REGION Network 10: Bit 9
   RUNG wire#powerrail
      Contact( #wInWord.%X9 )
      Coil( #bOutBit09 )
   END_RUNG
   // the same network as SCL:
   #bOutBit09 := #wInWord.%X9;
END_REGION

REGION Network 11: Bit 10
   RUNG wire#powerrail
      Contact( #wInWord.%X10 )
      Coil( #bOutBit10 )
   END_RUNG
   // the same network as SCL:
   #bOutBit10 := #wInWord.%X10;
END_REGION

REGION Network 12: Bit 11
   RUNG wire#powerrail
      Contact( #wInWord.%X11 )
      Coil( #bOutBit11 )
   END_RUNG
   // the same network as SCL:
   #bOutBit11 := #wInWord.%X11;
END_REGION

REGION Network 13: Bit 12
   RUNG wire#powerrail
      Contact( #wInWord.%X12 )
      Coil( #bOutBit12 )
   END_RUNG
   // the same network as SCL:
   #bOutBit12 := #wInWord.%X12;
END_REGION

REGION Network 14: Bit 13
   RUNG wire#powerrail
      Contact( #wInWord.%X13 )
      Coil( #bOutBit13 )
   END_RUNG
   // the same network as SCL:
   #bOutBit13 := #wInWord.%X13;
END_REGION

REGION Network 15: Bit 14
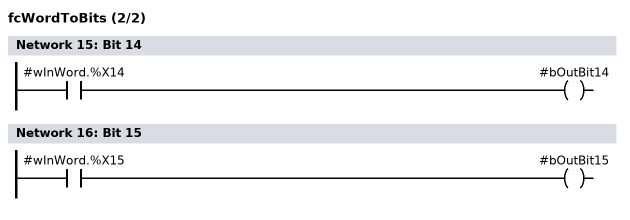
   RUNG wire#powerrail
      Contact( #wInWord.%X14 )
      Coil( #bOutBit14 )
   END_RUNG
   // the same network as SCL:
   #bOutBit14 := #wInWord.%X14;
END_REGION

REGION Network 16: Bit 15
   RUNG wire#powerrail
      Contact( #wInWord.%X15 )
      Coil( #bOutBit15 )
   END_RUNG
   // the same network as SCL:
   #bOutBit15 := #wInWord.%X15;
END_REGION
END_FUNCTION

FUNCTION "fcBitsToWord" : Void   // FC1001, LAD
TITLE = Pack Bits into word
{ S7_Optimized_Access := 'FALSE' }
AUTHOR : DMC
FAMILY : LowLevel
VERSION : 0.1
BEGIN

REGION Network 1: Bit0
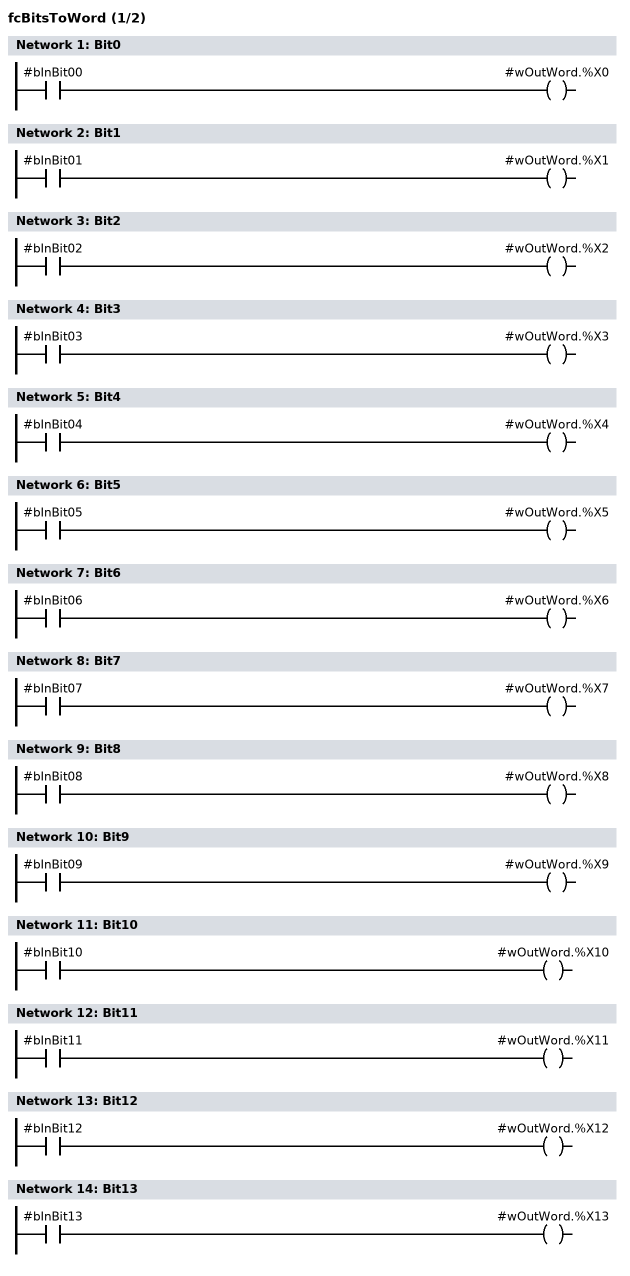
   RUNG wire#powerrail
      Contact( #bInBit00 )
      Coil( #wOutWord.%X0 )
   END_RUNG
   // the same network as SCL:
   #wOutWord.%X0 := #bInBit00;
END_REGION

REGION Network 2: Bit1
   RUNG wire#powerrail
      Contact( #bInBit01 )
      Coil( #wOutWord.%X1 )
   END_RUNG
   // the same network as SCL:
   #wOutWord.%X1 := #bInBit01;
END_REGION

REGION Network 3: Bit2
   RUNG wire#powerrail
      Contact( #bInBit02 )
      Coil( #wOutWord.%X2 )
   END_RUNG
   // the same network as SCL:
   #wOutWord.%X2 := #bInBit02;
END_REGION

REGION Network 4: Bit3
   RUNG wire#powerrail
      Contact( #bInBit03 )
      Coil( #wOutWord.%X3 )
   END_RUNG
   // the same network as SCL:
   #wOutWord.%X3 := #bInBit03;
END_REGION

REGION Network 5: Bit4
   RUNG wire#powerrail
      Contact( #bInBit04 )
      Coil( #wOutWord.%X4 )
   END_RUNG
   // the same network as SCL:
   #wOutWord.%X4 := #bInBit04;
END_REGION

REGION Network 6: Bit5
   RUNG wire#powerrail
      Contact( #bInBit05 )
      Coil( #wOutWord.%X5 )
   END_RUNG
   // the same network as SCL:
   #wOutWord.%X5 := #bInBit05;
END_REGION

REGION Network 7: Bit6
   RUNG wire#powerrail
      Contact( #bInBit06 )
      Coil( #wOutWord.%X6 )
   END_RUNG
   // the same network as SCL:
   #wOutWord.%X6 := #bInBit06;
END_REGION

REGION Network 8: Bit7
   RUNG wire#powerrail
      Contact( #bInBit07 )
      Coil( #wOutWord.%X7 )
   END_RUNG
   // the same network as SCL:
   #wOutWord.%X7 := #bInBit07;
END_REGION

REGION Network 9: Bit8
   RUNG wire#powerrail
      Contact( #bInBit08 )
      Coil( #wOutWord.%X8 )
   END_RUNG
   // the same network as SCL:
   #wOutWord.%X8 := #bInBit08;
END_REGION

REGION Network 10: Bit9
   RUNG wire#powerrail
      Contact( #bInBit09 )
      Coil( #wOutWord.%X9 )
   END_RUNG
   // the same network as SCL:
   #wOutWord.%X9 := #bInBit09;
END_REGION

REGION Network 11: Bit10
   RUNG wire#powerrail
      Contact( #bInBit10 )
      Coil( #wOutWord.%X10 )
   END_RUNG
   // the same network as SCL:
   #wOutWord.%X10 := #bInBit10;
END_REGION

REGION Network 12: Bit11
   RUNG wire#powerrail
      Contact( #bInBit11 )
      Coil( #wOutWord.%X11 )
   END_RUNG
   // the same network as SCL:
   #wOutWord.%X11 := #bInBit11;
END_REGION

REGION Network 13: Bit12
   RUNG wire#powerrail
      Contact( #bInBit12 )
      Coil( #wOutWord.%X12 )
   END_RUNG
   // the same network as SCL:
   #wOutWord.%X12 := #bInBit12;
END_REGION

REGION Network 14: Bit13
   RUNG wire#powerrail
      Contact( #bInBit13 )
      Coil( #wOutWord.%X13 )
   END_RUNG
   // the same network as SCL:
   #wOutWord.%X13 := #bInBit13;
END_REGION

REGION Network 15: Bit14
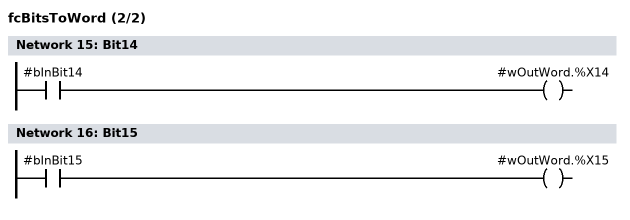
   RUNG wire#powerrail
      Contact( #bInBit14 )
      Coil( #wOutWord.%X14 )
   END_RUNG
   // the same network as SCL:
   #wOutWord.%X14 := #bInBit14;
END_REGION

REGION Network 16: Bit15
   RUNG wire#powerrail
      Contact( #bInBit15 )
      Coil( #wOutWord.%X15 )
   END_RUNG
   // the same network as SCL:
   #wOutWord.%X15 := #bInBit15;
END_REGION
END_FUNCTION

// folder: Library Blocks/Resources/HMI

FUNCTION_BLOCK "fbErrorScroller"   // FB1007, LAD
TITLE = Scrolls through the error codes for display on the HMI
{ S7_Optimized_Access := 'FALSE' }
AUTHOR : DMC
FAMILY : Error
VERSION : 0.1
   VAR_TEMP   // added for the SCL form of the ladder/FBD networks
      _w1 : Bool;
   END_VAR
BEGIN

REGION Network 1: Error Exists
   // OR all of the possible errors. If any error Exists, SET bErrorExists
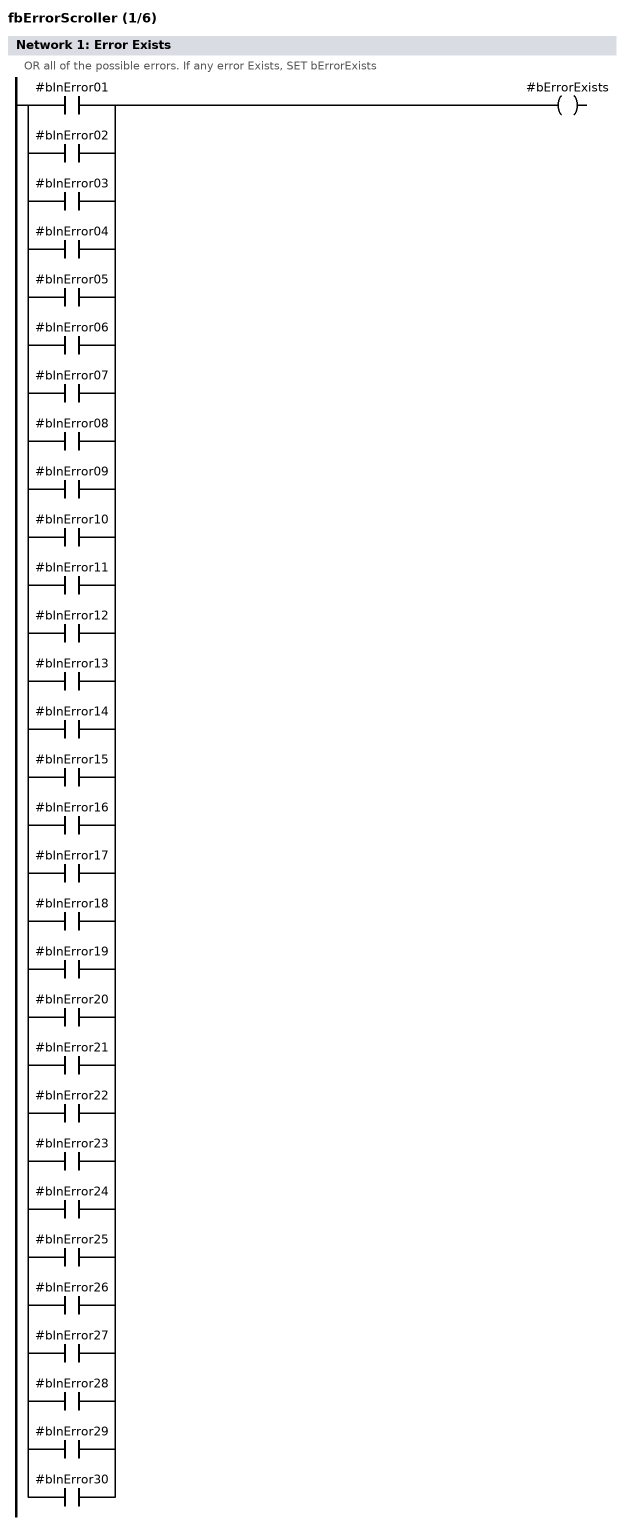
   RUNG wire#powerrail
      Contact( #bInError01 )
      wire#w1
      Coil( #bErrorExists )
   END_RUNG
   RUNG wire#powerrail
      Contact( #bInError02 )
   END_RUNG wire#w1
   RUNG wire#powerrail
      Contact( #bInError03 )
   END_RUNG wire#w1
   RUNG wire#powerrail
      Contact( #bInError04 )
   END_RUNG wire#w1
   RUNG wire#powerrail
      Contact( #bInError05 )
   END_RUNG wire#w1
   RUNG wire#powerrail
      Contact( #bInError06 )
   END_RUNG wire#w1
   RUNG wire#powerrail
      Contact( #bInError07 )
   END_RUNG wire#w1
   RUNG wire#powerrail
      Contact( #bInError08 )
   END_RUNG wire#w1
   RUNG wire#powerrail
      Contact( #bInError09 )
   END_RUNG wire#w1
   RUNG wire#powerrail
      Contact( #bInError10 )
   END_RUNG wire#w1
   RUNG wire#powerrail
      Contact( #bInError11 )
   END_RUNG wire#w1
   RUNG wire#powerrail
      Contact( #bInError12 )
   END_RUNG wire#w1
   RUNG wire#powerrail
      Contact( #bInError13 )
   END_RUNG wire#w1
   RUNG wire#powerrail
      Contact( #bInError14 )
   END_RUNG wire#w1
   RUNG wire#powerrail
      Contact( #bInError15 )
   END_RUNG wire#w1
   RUNG wire#powerrail
      Contact( #bInError16 )
   END_RUNG wire#w1
   RUNG wire#powerrail
      Contact( #bInError17 )
   END_RUNG wire#w1
   RUNG wire#powerrail
      Contact( #bInError18 )
   END_RUNG wire#w1
   RUNG wire#powerrail
      Contact( #bInError19 )
   END_RUNG wire#w1
   RUNG wire#powerrail
      Contact( #bInError20 )
   END_RUNG wire#w1
   RUNG wire#powerrail
      Contact( #bInError21 )
   END_RUNG wire#w1
   RUNG wire#powerrail
      Contact( #bInError22 )
   END_RUNG wire#w1
   RUNG wire#powerrail
      Contact( #bInError23 )
   END_RUNG wire#w1
   RUNG wire#powerrail
      Contact( #bInError24 )
   END_RUNG wire#w1
   RUNG wire#powerrail
      Contact( #bInError25 )
   END_RUNG wire#w1
   RUNG wire#powerrail
      Contact( #bInError26 )
   END_RUNG wire#w1
   RUNG wire#powerrail
      Contact( #bInError27 )
   END_RUNG wire#w1
   RUNG wire#powerrail
      Contact( #bInError28 )
   END_RUNG wire#w1
   RUNG wire#powerrail
      Contact( #bInError29 )
   END_RUNG wire#w1
   RUNG wire#powerrail
      Contact( #bInError30 )
   END_RUNG wire#w1
   // the same network as SCL:
   #bErrorExists := #bInError01 OR #bInError02 OR #bInError03 OR #bInError04 OR #bInError05 OR #bInError06 OR #bInError07 OR #bInError08 OR #bInError09 OR #bInError10 OR #bInError11 OR #bInError12 OR #bInError13 OR #bInError14 OR #bInError15 OR #bInError16 OR #bInError17 OR #bInError18 OR #bInError19 OR #bInError20 OR #bInError21 OR #bInError22 OR #bInError23 OR #bInError24 OR #bInError25 OR #bInError26 OR #bInError27 OR #bInError28 OR #bInError29 OR #bInError30;
END_REGION

REGION Network 2
   // ============================ Scroll errors on HMI ========================
   // Timed delay
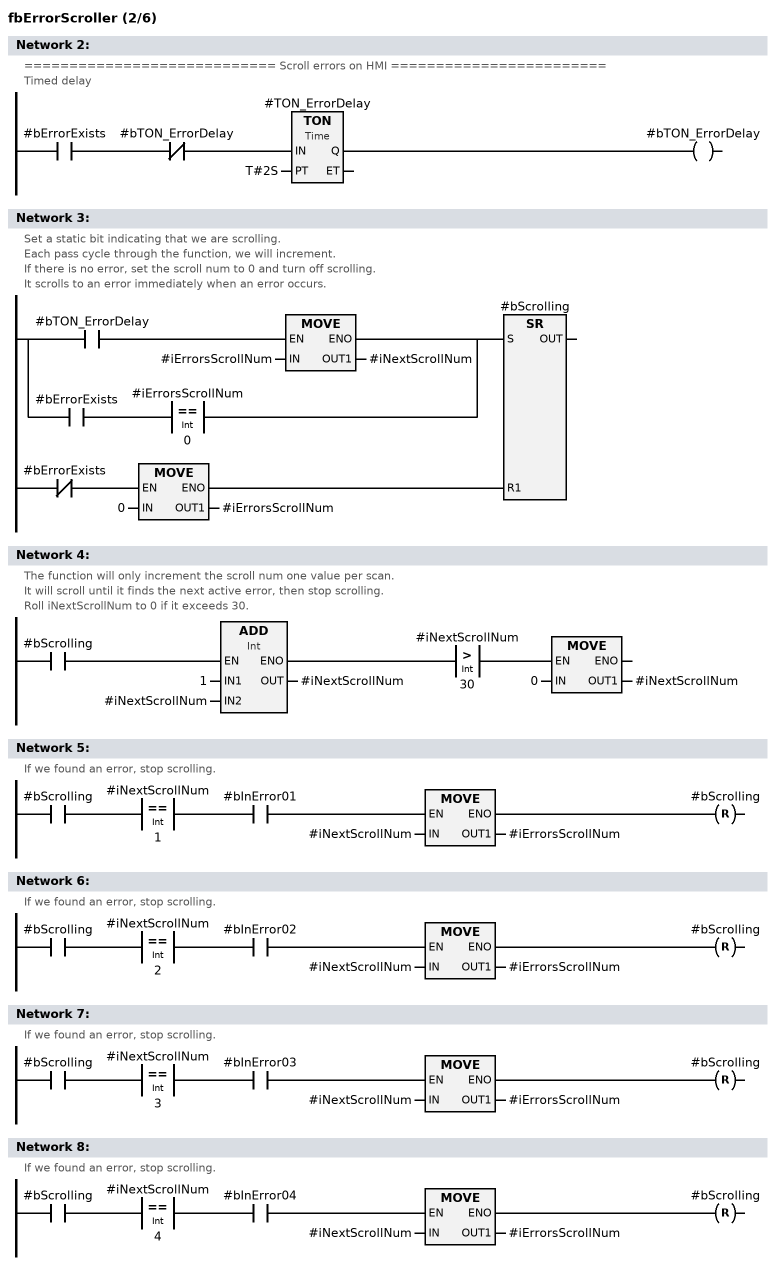
   #TON_ErrorDelay.TON(IN := #bErrorExists AND NOT #bTON_ErrorDelay, PT := T#2S);
   #bTON_ErrorDelay := #TON_ErrorDelay.Q;
END_REGION

REGION Network 3
   // Set a static bit indicating that we are scrolling.  
   // Each pass cycle through the function, we will increment.  
   // If there is no error, set the scroll num to 0 and turn off scrolling.  
   // It scrolls to an error immediately when an error occurs.
   RUNG wire#powerrail
      Contact( #bTON_ErrorDelay )
      { S7_GenerateENO := "TRUE" } Move(in := #iErrorsScrollNum, out1 => #iNextScrollNum)
      wire#w1
      S_SR(operand := #bScrolling, r1 := wire#w2)
   END_RUNG
   RUNG wire#powerrail
      Contact( #bErrorExists )
      { S7_Templates := "SrcType := Int" } EQ_Contact(in1 := #iErrorsScrollNum, in2 := 0)
   END_RUNG wire#w1
   RUNG wire#powerrail
      I_Contact( #bErrorExists )
      { S7_GenerateENO := "TRUE" } Move(in := 0, out1 => #iErrorsScrollNum)
   END_RUNG wire#w2
   // the same network as SCL:
   // ENO of a box is taken as its EN; it also drops when the box reports an error
   IF #bTON_ErrorDelay THEN #iNextScrollNum := #iErrorsScrollNum; END_IF;
   #_w1 := #bTON_ErrorDelay OR (#bErrorExists AND (#iErrorsScrollNum = 0));
   IF NOT #bErrorExists THEN #iErrorsScrollNum := 0; END_IF;
   IF #_w1 THEN
       #bScrolling := TRUE;   // SR flip-flop
   END_IF;
   IF NOT #bErrorExists THEN #bScrolling := FALSE; END_IF;
END_REGION

REGION Network 4
   // The function will only increment the scroll num one value per scan.  
   // It will scroll until it finds the next active error, then stop scrolling.  
   // Roll iNextScrollNum to 0 if it exceeds 30.
   RUNG wire#powerrail
      Contact( #bScrolling )
      { S7_Templates := "SrcType := Int"; S7_GenerateENO := "TRUE" } Add(in1 := 1, in2 := #iNextScrollNum, out => #iNextScrollNum)
      { S7_Templates := "SrcType := Int" } GT_Contact(in1 := #iNextScrollNum, in2 := 30)
      { S7_GenerateENO := "TRUE" } Move(in := 0, out1 => #iNextScrollNum)
   END_RUNG
   // the same network as SCL:
   // ENO of a box is taken as its EN; it also drops when the box reports an error
   IF #bScrolling THEN #iNextScrollNum := 1 + #iNextScrollNum; END_IF;
   IF #bScrolling AND (#iNextScrollNum > 30) THEN #iNextScrollNum := 0; END_IF;
END_REGION

REGION Network 5
   // If we found an error, stop scrolling.
   RUNG wire#powerrail
      Contact( #bScrolling )
      { S7_Templates := "SrcType := Int" } EQ_Contact(in1 := #iNextScrollNum, in2 := 1)
      Contact( #bInError01 )
      { S7_GenerateENO := "TRUE" } Move(in := #iNextScrollNum, out1 => #iErrorsScrollNum)
      R_Coil( #bScrolling )
   END_RUNG
   // the same network as SCL:
   // ENO of a box is taken as its EN; it also drops when the box reports an error
   IF #bScrolling AND (#iNextScrollNum = 1) AND #bInError01 THEN
       #iErrorsScrollNum := #iNextScrollNum;
       #bScrolling := FALSE;
   END_IF;
END_REGION

REGION Network 6
   // If we found an error, stop scrolling.
   RUNG wire#powerrail
      Contact( #bScrolling )
      { S7_Templates := "SrcType := Int" } EQ_Contact(in1 := #iNextScrollNum, in2 := 2)
      Contact( #bInError02 )
      { S7_GenerateENO := "TRUE" } Move(in := #iNextScrollNum, out1 => #iErrorsScrollNum)
      R_Coil( #bScrolling )
   END_RUNG
   // the same network as SCL:
   // ENO of a box is taken as its EN; it also drops when the box reports an error
   IF #bScrolling AND (#iNextScrollNum = 2) AND #bInError02 THEN
       #iErrorsScrollNum := #iNextScrollNum;
       #bScrolling := FALSE;
   END_IF;
END_REGION

REGION Network 7
   // If we found an error, stop scrolling.
   RUNG wire#powerrail
      Contact( #bScrolling )
      { S7_Templates := "SrcType := Int" } EQ_Contact(in1 := #iNextScrollNum, in2 := 3)
      Contact( #bInError03 )
      { S7_GenerateENO := "TRUE" } Move(in := #iNextScrollNum, out1 => #iErrorsScrollNum)
      R_Coil( #bScrolling )
   END_RUNG
   // the same network as SCL:
   // ENO of a box is taken as its EN; it also drops when the box reports an error
   IF #bScrolling AND (#iNextScrollNum = 3) AND #bInError03 THEN
       #iErrorsScrollNum := #iNextScrollNum;
       #bScrolling := FALSE;
   END_IF;
END_REGION

REGION Network 8
   // If we found an error, stop scrolling.
   RUNG wire#powerrail
      Contact( #bScrolling )
      { S7_Templates := "SrcType := Int" } EQ_Contact(in1 := #iNextScrollNum, in2 := 4)
      Contact( #bInError04 )
      { S7_GenerateENO := "TRUE" } Move(in := #iNextScrollNum, out1 => #iErrorsScrollNum)
      R_Coil( #bScrolling )
   END_RUNG
   // the same network as SCL:
   // ENO of a box is taken as its EN; it also drops when the box reports an error
   IF #bScrolling AND (#iNextScrollNum = 4) AND #bInError04 THEN
       #iErrorsScrollNum := #iNextScrollNum;
       #bScrolling := FALSE;
   END_IF;
END_REGION

REGION Network 9
   // If we found an error, stop scrolling.
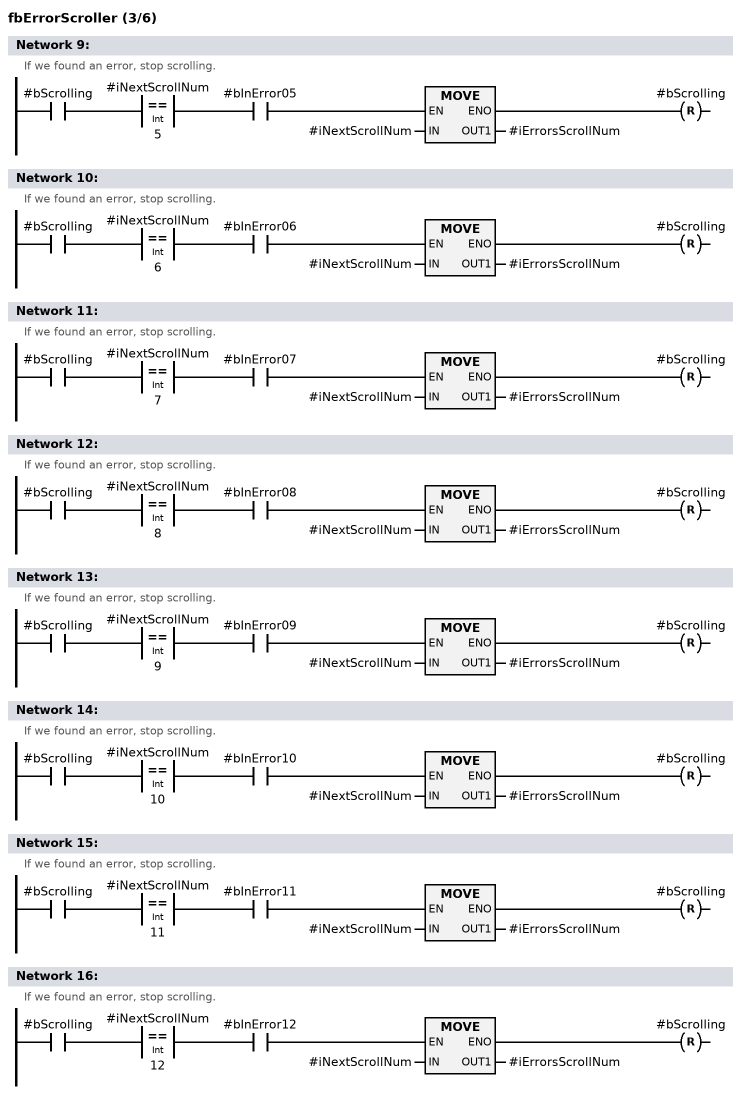
   RUNG wire#powerrail
      Contact( #bScrolling )
      { S7_Templates := "SrcType := Int" } EQ_Contact(in1 := #iNextScrollNum, in2 := 5)
      Contact( #bInError05 )
      { S7_GenerateENO := "TRUE" } Move(in := #iNextScrollNum, out1 => #iErrorsScrollNum)
      R_Coil( #bScrolling )
   END_RUNG
   // the same network as SCL:
   // ENO of a box is taken as its EN; it also drops when the box reports an error
   IF #bScrolling AND (#iNextScrollNum = 5) AND #bInError05 THEN
       #iErrorsScrollNum := #iNextScrollNum;
       #bScrolling := FALSE;
   END_IF;
END_REGION

REGION Network 10
   // If we found an error, stop scrolling.
   RUNG wire#powerrail
      Contact( #bScrolling )
      { S7_Templates := "SrcType := Int" } EQ_Contact(in1 := #iNextScrollNum, in2 := 6)
      Contact( #bInError06 )
      { S7_GenerateENO := "TRUE" } Move(in := #iNextScrollNum, out1 => #iErrorsScrollNum)
      R_Coil( #bScrolling )
   END_RUNG
   // the same network as SCL:
   // ENO of a box is taken as its EN; it also drops when the box reports an error
   IF #bScrolling AND (#iNextScrollNum = 6) AND #bInError06 THEN
       #iErrorsScrollNum := #iNextScrollNum;
       #bScrolling := FALSE;
   END_IF;
END_REGION

REGION Network 11
   // If we found an error, stop scrolling.
   RUNG wire#powerrail
      Contact( #bScrolling )
      { S7_Templates := "SrcType := Int" } EQ_Contact(in1 := #iNextScrollNum, in2 := 7)
      Contact( #bInError07 )
      { S7_GenerateENO := "TRUE" } Move(in := #iNextScrollNum, out1 => #iErrorsScrollNum)
      R_Coil( #bScrolling )
   END_RUNG
   // the same network as SCL:
   // ENO of a box is taken as its EN; it also drops when the box reports an error
   IF #bScrolling AND (#iNextScrollNum = 7) AND #bInError07 THEN
       #iErrorsScrollNum := #iNextScrollNum;
       #bScrolling := FALSE;
   END_IF;
END_REGION

REGION Network 12
   // If we found an error, stop scrolling.
   RUNG wire#powerrail
      Contact( #bScrolling )
      { S7_Templates := "SrcType := Int" } EQ_Contact(in1 := #iNextScrollNum, in2 := 8)
      Contact( #bInError08 )
      { S7_GenerateENO := "TRUE" } Move(in := #iNextScrollNum, out1 => #iErrorsScrollNum)
      R_Coil( #bScrolling )
   END_RUNG
   // the same network as SCL:
   // ENO of a box is taken as its EN; it also drops when the box reports an error
   IF #bScrolling AND (#iNextScrollNum = 8) AND #bInError08 THEN
       #iErrorsScrollNum := #iNextScrollNum;
       #bScrolling := FALSE;
   END_IF;
END_REGION

REGION Network 13
   // If we found an error, stop scrolling.
   RUNG wire#powerrail
      Contact( #bScrolling )
      { S7_Templates := "SrcType := Int" } EQ_Contact(in1 := #iNextScrollNum, in2 := 9)
      Contact( #bInError09 )
      { S7_GenerateENO := "TRUE" } Move(in := #iNextScrollNum, out1 => #iErrorsScrollNum)
      R_Coil( #bScrolling )
   END_RUNG
   // the same network as SCL:
   // ENO of a box is taken as its EN; it also drops when the box reports an error
   IF #bScrolling AND (#iNextScrollNum = 9) AND #bInError09 THEN
       #iErrorsScrollNum := #iNextScrollNum;
       #bScrolling := FALSE;
   END_IF;
END_REGION

REGION Network 14
   // If we found an error, stop scrolling.
   RUNG wire#powerrail
      Contact( #bScrolling )
      { S7_Templates := "SrcType := Int" } EQ_Contact(in1 := #iNextScrollNum, in2 := 10)
      Contact( #bInError10 )
      { S7_GenerateENO := "TRUE" } Move(in := #iNextScrollNum, out1 => #iErrorsScrollNum)
      R_Coil( #bScrolling )
   END_RUNG
   // the same network as SCL:
   // ENO of a box is taken as its EN; it also drops when the box reports an error
   IF #bScrolling AND (#iNextScrollNum = 10) AND #bInError10 THEN
       #iErrorsScrollNum := #iNextScrollNum;
       #bScrolling := FALSE;
   END_IF;
END_REGION

REGION Network 15
   // If we found an error, stop scrolling.
   RUNG wire#powerrail
      Contact( #bScrolling )
      { S7_Templates := "SrcType := Int" } EQ_Contact(in1 := #iNextScrollNum, in2 := 11)
      Contact( #bInError11 )
      { S7_GenerateENO := "TRUE" } Move(in := #iNextScrollNum, out1 => #iErrorsScrollNum)
      R_Coil( #bScrolling )
   END_RUNG
   // the same network as SCL:
   // ENO of a box is taken as its EN; it also drops when the box reports an error
   IF #bScrolling AND (#iNextScrollNum = 11) AND #bInError11 THEN
       #iErrorsScrollNum := #iNextScrollNum;
       #bScrolling := FALSE;
   END_IF;
END_REGION

REGION Network 16
   // If we found an error, stop scrolling.
   RUNG wire#powerrail
      Contact( #bScrolling )
      { S7_Templates := "SrcType := Int" } EQ_Contact(in1 := #iNextScrollNum, in2 := 12)
      Contact( #bInError12 )
      { S7_GenerateENO := "TRUE" } Move(in := #iNextScrollNum, out1 => #iErrorsScrollNum)
      R_Coil( #bScrolling )
   END_RUNG
   // the same network as SCL:
   // ENO of a box is taken as its EN; it also drops when the box reports an error
   IF #bScrolling AND (#iNextScrollNum = 12) AND #bInError12 THEN
       #iErrorsScrollNum := #iNextScrollNum;
       #bScrolling := FALSE;
   END_IF;
END_REGION

REGION Network 17
   // If we found an error, stop scrolling.
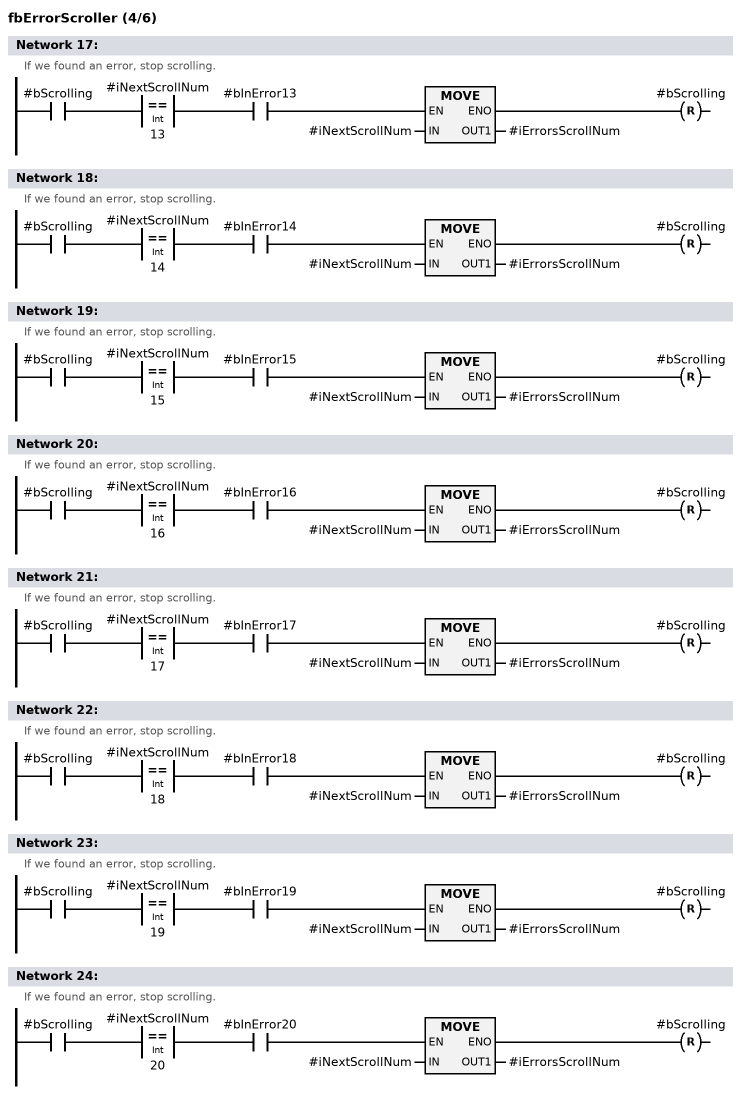
   RUNG wire#powerrail
      Contact( #bScrolling )
      { S7_Templates := "SrcType := Int" } EQ_Contact(in1 := #iNextScrollNum, in2 := 13)
      Contact( #bInError13 )
      { S7_GenerateENO := "TRUE" } Move(in := #iNextScrollNum, out1 => #iErrorsScrollNum)
      R_Coil( #bScrolling )
   END_RUNG
   // the same network as SCL:
   // ENO of a box is taken as its EN; it also drops when the box reports an error
   IF #bScrolling AND (#iNextScrollNum = 13) AND #bInError13 THEN
       #iErrorsScrollNum := #iNextScrollNum;
       #bScrolling := FALSE;
   END_IF;
END_REGION

REGION Network 18
   // If we found an error, stop scrolling.
   RUNG wire#powerrail
      Contact( #bScrolling )
      { S7_Templates := "SrcType := Int" } EQ_Contact(in1 := #iNextScrollNum, in2 := 14)
      Contact( #bInError14 )
      { S7_GenerateENO := "TRUE" } Move(in := #iNextScrollNum, out1 => #iErrorsScrollNum)
      R_Coil( #bScrolling )
   END_RUNG
   // the same network as SCL:
   // ENO of a box is taken as its EN; it also drops when the box reports an error
   IF #bScrolling AND (#iNextScrollNum = 14) AND #bInError14 THEN
       #iErrorsScrollNum := #iNextScrollNum;
       #bScrolling := FALSE;
   END_IF;
END_REGION

REGION Network 19
   // If we found an error, stop scrolling.
   RUNG wire#powerrail
      Contact( #bScrolling )
      { S7_Templates := "SrcType := Int" } EQ_Contact(in1 := #iNextScrollNum, in2 := 15)
      Contact( #bInError15 )
      { S7_GenerateENO := "TRUE" } Move(in := #iNextScrollNum, out1 => #iErrorsScrollNum)
      R_Coil( #bScrolling )
   END_RUNG
   // the same network as SCL:
   // ENO of a box is taken as its EN; it also drops when the box reports an error
   IF #bScrolling AND (#iNextScrollNum = 15) AND #bInError15 THEN
       #iErrorsScrollNum := #iNextScrollNum;
       #bScrolling := FALSE;
   END_IF;
END_REGION

REGION Network 20
   // If we found an error, stop scrolling.
   RUNG wire#powerrail
      Contact( #bScrolling )
      { S7_Templates := "SrcType := Int" } EQ_Contact(in1 := #iNextScrollNum, in2 := 16)
      Contact( #bInError16 )
      { S7_GenerateENO := "TRUE" } Move(in := #iNextScrollNum, out1 => #iErrorsScrollNum)
      R_Coil( #bScrolling )
   END_RUNG
   // the same network as SCL:
   // ENO of a box is taken as its EN; it also drops when the box reports an error
   IF #bScrolling AND (#iNextScrollNum = 16) AND #bInError16 THEN
       #iErrorsScrollNum := #iNextScrollNum;
       #bScrolling := FALSE;
   END_IF;
END_REGION

REGION Network 21
   // If we found an error, stop scrolling.
   RUNG wire#powerrail
      Contact( #bScrolling )
      { S7_Templates := "SrcType := Int" } EQ_Contact(in1 := #iNextScrollNum, in2 := 17)
      Contact( #bInError17 )
      { S7_GenerateENO := "TRUE" } Move(in := #iNextScrollNum, out1 => #iErrorsScrollNum)
      R_Coil( #bScrolling )
   END_RUNG
   // the same network as SCL:
   // ENO of a box is taken as its EN; it also drops when the box reports an error
   IF #bScrolling AND (#iNextScrollNum = 17) AND #bInError17 THEN
       #iErrorsScrollNum := #iNextScrollNum;
       #bScrolling := FALSE;
   END_IF;
END_REGION

REGION Network 22
   // If we found an error, stop scrolling.
   RUNG wire#powerrail
      Contact( #bScrolling )
      { S7_Templates := "SrcType := Int" } EQ_Contact(in1 := #iNextScrollNum, in2 := 18)
      Contact( #bInError18 )
      { S7_GenerateENO := "TRUE" } Move(in := #iNextScrollNum, out1 => #iErrorsScrollNum)
      R_Coil( #bScrolling )
   END_RUNG
   // the same network as SCL:
   // ENO of a box is taken as its EN; it also drops when the box reports an error
   IF #bScrolling AND (#iNextScrollNum = 18) AND #bInError18 THEN
       #iErrorsScrollNum := #iNextScrollNum;
       #bScrolling := FALSE;
   END_IF;
END_REGION

REGION Network 23
   // If we found an error, stop scrolling.
   RUNG wire#powerrail
      Contact( #bScrolling )
      { S7_Templates := "SrcType := Int" } EQ_Contact(in1 := #iNextScrollNum, in2 := 19)
      Contact( #bInError19 )
      { S7_GenerateENO := "TRUE" } Move(in := #iNextScrollNum, out1 => #iErrorsScrollNum)
      R_Coil( #bScrolling )
   END_RUNG
   // the same network as SCL:
   // ENO of a box is taken as its EN; it also drops when the box reports an error
   IF #bScrolling AND (#iNextScrollNum = 19) AND #bInError19 THEN
       #iErrorsScrollNum := #iNextScrollNum;
       #bScrolling := FALSE;
   END_IF;
END_REGION

REGION Network 24
   // If we found an error, stop scrolling.
   RUNG wire#powerrail
      Contact( #bScrolling )
      { S7_Templates := "SrcType := Int" } EQ_Contact(in1 := #iNextScrollNum, in2 := 20)
      Contact( #bInError20 )
      { S7_GenerateENO := "TRUE" } Move(in := #iNextScrollNum, out1 => #iErrorsScrollNum)
      R_Coil( #bScrolling )
   END_RUNG
   // the same network as SCL:
   // ENO of a box is taken as its EN; it also drops when the box reports an error
   IF #bScrolling AND (#iNextScrollNum = 20) AND #bInError20 THEN
       #iErrorsScrollNum := #iNextScrollNum;
       #bScrolling := FALSE;
   END_IF;
END_REGION

REGION Network 25
   // If we found an error, stop scrolling.
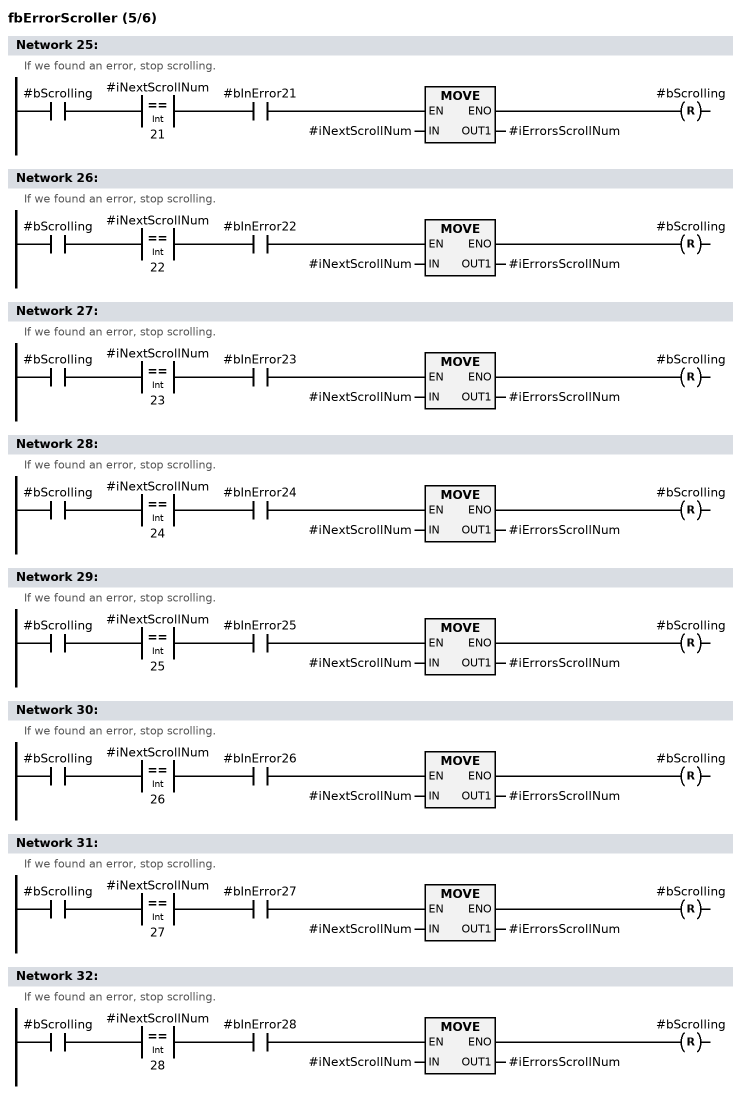
   RUNG wire#powerrail
      Contact( #bScrolling )
      { S7_Templates := "SrcType := Int" } EQ_Contact(in1 := #iNextScrollNum, in2 := 21)
      Contact( #bInError21 )
      { S7_GenerateENO := "TRUE" } Move(in := #iNextScrollNum, out1 => #iErrorsScrollNum)
      R_Coil( #bScrolling )
   END_RUNG
   // the same network as SCL:
   // ENO of a box is taken as its EN; it also drops when the box reports an error
   IF #bScrolling AND (#iNextScrollNum = 21) AND #bInError21 THEN
       #iErrorsScrollNum := #iNextScrollNum;
       #bScrolling := FALSE;
   END_IF;
END_REGION

REGION Network 26
   // If we found an error, stop scrolling.
   RUNG wire#powerrail
      Contact( #bScrolling )
      { S7_Templates := "SrcType := Int" } EQ_Contact(in1 := #iNextScrollNum, in2 := 22)
      Contact( #bInError22 )
      { S7_GenerateENO := "TRUE" } Move(in := #iNextScrollNum, out1 => #iErrorsScrollNum)
      R_Coil( #bScrolling )
   END_RUNG
   // the same network as SCL:
   // ENO of a box is taken as its EN; it also drops when the box reports an error
   IF #bScrolling AND (#iNextScrollNum = 22) AND #bInError22 THEN
       #iErrorsScrollNum := #iNextScrollNum;
       #bScrolling := FALSE;
   END_IF;
END_REGION

REGION Network 27
   // If we found an error, stop scrolling.
   RUNG wire#powerrail
      Contact( #bScrolling )
      { S7_Templates := "SrcType := Int" } EQ_Contact(in1 := #iNextScrollNum, in2 := 23)
      Contact( #bInError23 )
      { S7_GenerateENO := "TRUE" } Move(in := #iNextScrollNum, out1 => #iErrorsScrollNum)
      R_Coil( #bScrolling )
   END_RUNG
   // the same network as SCL:
   // ENO of a box is taken as its EN; it also drops when the box reports an error
   IF #bScrolling AND (#iNextScrollNum = 23) AND #bInError23 THEN
       #iErrorsScrollNum := #iNextScrollNum;
       #bScrolling := FALSE;
   END_IF;
END_REGION

REGION Network 28
   // If we found an error, stop scrolling.
   RUNG wire#powerrail
      Contact( #bScrolling )
      { S7_Templates := "SrcType := Int" } EQ_Contact(in1 := #iNextScrollNum, in2 := 24)
      Contact( #bInError24 )
      { S7_GenerateENO := "TRUE" } Move(in := #iNextScrollNum, out1 => #iErrorsScrollNum)
      R_Coil( #bScrolling )
   END_RUNG
   // the same network as SCL:
   // ENO of a box is taken as its EN; it also drops when the box reports an error
   IF #bScrolling AND (#iNextScrollNum = 24) AND #bInError24 THEN
       #iErrorsScrollNum := #iNextScrollNum;
       #bScrolling := FALSE;
   END_IF;
END_REGION

REGION Network 29
   // If we found an error, stop scrolling.
   RUNG wire#powerrail
      Contact( #bScrolling )
      { S7_Templates := "SrcType := Int" } EQ_Contact(in1 := #iNextScrollNum, in2 := 25)
      Contact( #bInError25 )
      { S7_GenerateENO := "TRUE" } Move(in := #iNextScrollNum, out1 => #iErrorsScrollNum)
      R_Coil( #bScrolling )
   END_RUNG
   // the same network as SCL:
   // ENO of a box is taken as its EN; it also drops when the box reports an error
   IF #bScrolling AND (#iNextScrollNum = 25) AND #bInError25 THEN
       #iErrorsScrollNum := #iNextScrollNum;
       #bScrolling := FALSE;
   END_IF;
END_REGION

REGION Network 30
   // If we found an error, stop scrolling.
   RUNG wire#powerrail
      Contact( #bScrolling )
      { S7_Templates := "SrcType := Int" } EQ_Contact(in1 := #iNextScrollNum, in2 := 26)
      Contact( #bInError26 )
      { S7_GenerateENO := "TRUE" } Move(in := #iNextScrollNum, out1 => #iErrorsScrollNum)
      R_Coil( #bScrolling )
   END_RUNG
   // the same network as SCL:
   // ENO of a box is taken as its EN; it also drops when the box reports an error
   IF #bScrolling AND (#iNextScrollNum = 26) AND #bInError26 THEN
       #iErrorsScrollNum := #iNextScrollNum;
       #bScrolling := FALSE;
   END_IF;
END_REGION

REGION Network 31
   // If we found an error, stop scrolling.
   RUNG wire#powerrail
      Contact( #bScrolling )
      { S7_Templates := "SrcType := Int" } EQ_Contact(in1 := #iNextScrollNum, in2 := 27)
      Contact( #bInError27 )
      { S7_GenerateENO := "TRUE" } Move(in := #iNextScrollNum, out1 => #iErrorsScrollNum)
      R_Coil( #bScrolling )
   END_RUNG
   // the same network as SCL:
   // ENO of a box is taken as its EN; it also drops when the box reports an error
   IF #bScrolling AND (#iNextScrollNum = 27) AND #bInError27 THEN
       #iErrorsScrollNum := #iNextScrollNum;
       #bScrolling := FALSE;
   END_IF;
END_REGION

REGION Network 32
   // If we found an error, stop scrolling.
   RUNG wire#powerrail
      Contact( #bScrolling )
      { S7_Templates := "SrcType := Int" } EQ_Contact(in1 := #iNextScrollNum, in2 := 28)
      Contact( #bInError28 )
      { S7_GenerateENO := "TRUE" } Move(in := #iNextScrollNum, out1 => #iErrorsScrollNum)
      R_Coil( #bScrolling )
   END_RUNG
   // the same network as SCL:
   // ENO of a box is taken as its EN; it also drops when the box reports an error
   IF #bScrolling AND (#iNextScrollNum = 28) AND #bInError28 THEN
       #iErrorsScrollNum := #iNextScrollNum;
       #bScrolling := FALSE;
   END_IF;
END_REGION

REGION Network 33
   // If we found an error, stop scrolling.
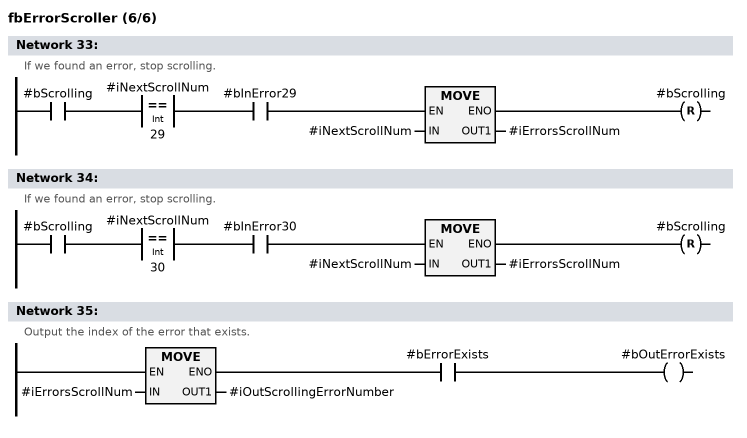
   RUNG wire#powerrail
      Contact( #bScrolling )
      { S7_Templates := "SrcType := Int" } EQ_Contact(in1 := #iNextScrollNum, in2 := 29)
      Contact( #bInError29 )
      { S7_GenerateENO := "TRUE" } Move(in := #iNextScrollNum, out1 => #iErrorsScrollNum)
      R_Coil( #bScrolling )
   END_RUNG
   // the same network as SCL:
   // ENO of a box is taken as its EN; it also drops when the box reports an error
   IF #bScrolling AND (#iNextScrollNum = 29) AND #bInError29 THEN
       #iErrorsScrollNum := #iNextScrollNum;
       #bScrolling := FALSE;
   END_IF;
END_REGION

REGION Network 34
   // If we found an error, stop scrolling.
   RUNG wire#powerrail
      Contact( #bScrolling )
      { S7_Templates := "SrcType := Int" } EQ_Contact(in1 := #iNextScrollNum, in2 := 30)
      Contact( #bInError30 )
      { S7_GenerateENO := "TRUE" } Move(in := #iNextScrollNum, out1 => #iErrorsScrollNum)
      R_Coil( #bScrolling )
   END_RUNG
   // the same network as SCL:
   // ENO of a box is taken as its EN; it also drops when the box reports an error
   IF #bScrolling AND (#iNextScrollNum = 30) AND #bInError30 THEN
       #iErrorsScrollNum := #iNextScrollNum;
       #bScrolling := FALSE;
   END_IF;
END_REGION

REGION Network 35
   // Output the index of the error that exists.
   RUNG wire#powerrail
      { S7_GenerateENO := "TRUE" } Move(in := #iErrorsScrollNum, out1 => #iOutScrollingErrorNumber)
      Contact( #bErrorExists )
      Coil( #bOutErrorExists )
   END_RUNG
   // the same network as SCL:
   // ENO of a box is taken as its EN; it also drops when the box reports an error
   #iOutScrollingErrorNumber := #iErrorsScrollNum;
   #bOutErrorExists := #bErrorExists;
END_REGION
END_FUNCTION_BLOCK

FUNCTION "fcHMIBit" : Void   // FC1030, LAD
{ S7_Optimized_Access := 'FALSE' }
VERSION : 0.1
   VAR_TEMP   // added for the SCL form of the ladder/FBD networks
      _w1 : Bool;
   END_VAR
BEGIN

REGION Network 1
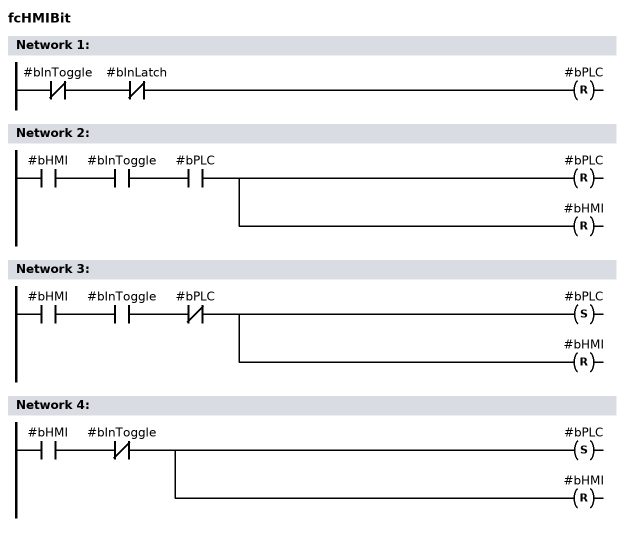
   RUNG wire#powerrail
      I_Contact( #bInToggle )
      I_Contact( #bInLatch )
      R_Coil( #bPLC )
   END_RUNG
   // the same network as SCL:
   IF NOT #bInToggle AND NOT #bInLatch THEN #bPLC := FALSE; END_IF;
END_REGION

REGION Network 2
   RUNG wire#powerrail
      Contact( #bHMI )
      Contact( #bInToggle )
      Contact( #bPLC )
      wire#w1
      R_Coil( #bPLC )
   END_RUNG
   RUNG wire#w1
      R_Coil( #bHMI )
   END_RUNG
   // the same network as SCL:
   #_w1 := #bHMI AND #bInToggle AND #bPLC;
   IF #_w1 THEN
       #bPLC := FALSE;
       #bHMI := FALSE;
   END_IF;
END_REGION

REGION Network 3
   RUNG wire#powerrail
      Contact( #bHMI )
      Contact( #bInToggle )
      I_Contact( #bPLC )
      wire#w1
      S_Coil( #bPLC )
   END_RUNG
   RUNG wire#w1
      R_Coil( #bHMI )
   END_RUNG
   // the same network as SCL:
   #_w1 := #bHMI AND #bInToggle AND NOT #bPLC;
   IF #_w1 THEN
       #bPLC := TRUE;
       #bHMI := FALSE;
   END_IF;
END_REGION

REGION Network 4
   RUNG wire#powerrail
      Contact( #bHMI )
      I_Contact( #bInToggle )
      wire#w1
      S_Coil( #bPLC )
   END_RUNG
   RUNG wire#w1
      R_Coil( #bHMI )
   END_RUNG
   // the same network as SCL:
   IF #bHMI AND NOT #bInToggle THEN
       #bPLC := TRUE;
       #bHMI := FALSE;
   END_IF;
END_REGION
END_FUNCTION

FUNCTION "fcSetHMIStatus" : Void   // FC1120, LAD
TITLE = Sets HMI Status
{ S7_Optimized_Access := 'FALSE' }
VERSION : 0.1
// Wrapper function for setting the HMI status of a device
// 
// In order of priority:
// 1. E-stop
// 2. Error
// 3. Forward/Work Position
// 4. Reverse/Home Position
// 5. Forward/Work On
// 6. Reverse/Home On
// 7. None
BEGIN

REGION Network 1: Set Reverse/Home On
